// TIA Portal project "opc_pc-station" (V16)

(* hardware
DEVICE "S7-1200 station_1"  S7-1200 Station
   slot 0: "Rack_0"  S7-1200 Rack  Rack  V1.0
   slot 1: "1214dc"  CPU 1214C DC/DC/DC  6ES7 214-1AG40-0XB0  V4.4
DEVICE "PC station"  SIMATIC PC station
   slot 0: "PC station"  Rail  SIMATIC PC-Station  V1.0
      slot 125: "Stationmanager"  Station_Manager  V6.0.4
   slot 1: "IE general_1"  IE General  IE_CP  V8.2.0
   slot 2: "OPC Server_1"  OPC Server  OPC Server  V16.0.0
DEVICE "S7300/ET200M station_1"  S7-300 station
   slot 0: "Rail_0"  Rail  6ES7 390-1***0-0AA0
   slot 2: "314c"  CPU 314C-2 PN/DP  6ES7 314-6EH04-0AB0  V3.3
      slot 2: "PROFINET interface_1"  PN-IO
         slot 1: "Port_1"  Port
         slot 2: "Port_2"  Port
      slot 5: "DI 24/DO 16_1"  DI24/DO16
      slot 6: "AI 5/AO 2_1"  AI5/AO2
      slot 7: "Count_1"  Counter
      slot 8: "Positioning_1"  Positioning
DEVICE "S71500/ET200MP station_1"  S7-1500 station
   slot 0: "Rail_0"  Rack  6ES7 590-1***0-0AA0
   slot 1: "1511f"  CPU 1511F-1 PN  6ES7 511-1FK02-0AB0  V2.8
      slot 3: "CPU display_1"  6ES7591-1AA00-0AA0
      slot 32768: "1511f"  X1
         slot 32769: "Port_1"  X1 P1
         slot 32770: "Port_2"  X1 P2
      slot 34817: "Virtual CP interface port_1"  Virtual CP interface port  Virtual CP interface port
DEVICE "S7300/ET200M station_2"  S7-300 station
   slot 0: "Rail_0"  Rail  6ES7 390-1***0-0AA0
   slot 2: "314c_cp343"  CPU 314C-2 PN/DP  6ES7 314-6EH04-0AB0  V3.3
      slot 2: "PROFINET interface_1"  PN-IO
         slot 1: "Port_1"  Port
         slot 2: "Port_2"  Port
      slot 5: "DI 24/DO 16_1"  DI24/DO16
      slot 6: "AI 5/AO 2_1"  AI5/AO2
      slot 7: "Count_1"  Counter
      slot 8: "Positioning_1"  Positioning
   slot 4: "CP 343-1 Advanced-IT_1"  CP 343-1 ADVANCED-IT  6GK7 343-1GX31-0XE0  V3.0
DEVICE "S71500/ET200MP station_2"  S7-1500 station
   slot 0: "Rail_0"  Rack  6ES7 590-1***0-0AA0
   slot 1: "1511f_cp"  CPU 1511F-1 PN  6ES7 511-1FK02-0AB0  V2.8
      slot 3: "CPU display_1"  6ES7591-1AA00-0AA0
      slot 32768: "1511f"  X1
         slot 32769: "Port_1"  X1 P1
         slot 32770: "Port_2"  X1 P2
      slot 34817: "Virtual CP interface port_1"  Virtual CP interface port  Virtual CP interface port
   slot 2: "CP 1543-1_1"  CP 1543-1  6GK7 543-1AX00-0XE0  V2.2
DEVICE "S7-1200 station_2"  S7-1200 Station
   slot 0: "Rack_0"  S7-1200 Rack  Rack  V1.0
   slot 1: "1212fc_cp"  CPU 1212FC DC/DC/DC  6ES7 212-1AF40-0XB0  V4.4
   slot 101: "CP 1243-1"  CP 1243-1  6GK7 243-1BX30-0XE0  V3.2
      slot 0: "Telecontrol server"  Partner
      slot 0: "Inter-station communication"  Partner
*)

// ===== PLC "1214dc"  CPU 1214C DC/DC/DC =====

VAR_GLOBAL   // PLC tag table "Default tag table"
   "Tag_clock" AT %MW2 : Int;
   "Tag_Int" AT %MW4 : Int;
END_VAR

DATA_BLOCK "data_db"   // DB1
{ S7_Optimized_Access := 'TRUE' }
VERSION : 0.1
   VAR
      zm_array : Array[0..2] of Byte;
      zm_bool : Bool;
      zm_byte : Byte;
      zm_char : Char;
      zm_datetime_dtl : DTL;
      zm_dword : DWord;
      zm_int : Int;
      zm_real : Real;
      zm_string : String;
      zm_struct : Struct
         zm_struct_bool : Bool;
         zm_struct_byte : Byte;
      END_STRUCT;
   END_VAR
BEGIN
END_DATA_BLOCK

ORGANIZATION_BLOCK "Main"   // OB1, LAD, ProgramCycle
TITLE = "Main Program Sweep (Cycle)"
{ S7_Optimized_Access := 'TRUE' }
VERSION : 0.1
   VAR_INPUT
      Initial_Call : Bool;   // Initial call of this OB
      Remanence : Bool;   // =True, if remanent data are available
   END_VAR
BEGIN

REGION Network 1
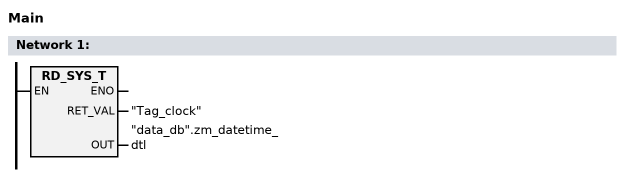
   "Tag_clock" := RD_SYS_T(OUT => "data_db".zm_datetime_dtl);
END_REGION
END_ORGANIZATION_BLOCK

// ===== PLC "314c"  CPU 314C-2 PN/DP =====

VAR_GLOBAL   // PLC tag table "Default tag table"
   "Tag_1" AT %MW0 : Int;
   "Tag_2" AT %M3.0 : Bool;
   "Tag_3" AT %MW4 : Word;
END_VAR

DATA_BLOCK "db_opc"   // DB1
{ S7_Optimized_Access := 'FALSE' }
VERSION : 0.1
   VAR
      zm_array : Array[0..2] of Byte;
      zm_bool : Bool;
      zm_byte : Byte;
      zm_char : Char;
      zm_datetime_rd_sys_t : Date_And_Time;
      zm_dword : DWord;
      zm_int : Int;
      zm_real : Real;
      zm_string : String;
      zm_struct : Struct
         zm_struct_bool : Bool;
         zm_struct_byte : Byte;
      END_STRUCT;
   END_VAR
BEGIN
END_DATA_BLOCK

ORGANIZATION_BLOCK "Main"   // OB1, LAD
TITLE = "Main Program Sweep (Cycle)"
{ S7_Optimized_Access := 'FALSE' }
VERSION : 0.1
   VAR_TEMP
      OB1_EV_CLASS : Byte;   // Bits 0-3 = 1 (Coming event), Bits 4-7 = 1 (Event class 1)
      OB1_SCAN_1 : Byte;   // 1 (Cold restart scan 1 of OB 1), 3 (Scan 2-n of OB 1)
      OB1_PRIORITY : Byte;   // Priority of OB Execution
      OB1_OB_NUMBR : Byte;   // 1 (Organization block 1, OB1)
      OB1_RESERVED_1 : Byte;   // Reserved for system
      OB1_RESERVED_2 : Byte;   // Reserved for system
      OB1_PREV_CYCLE : Int;   // Cycle time of previous OB1 scan (milliseconds)
      OB1_MIN_CYCLE : Int;   // Minimum cycle time of OB1 (milliseconds)
      OB1_MAX_CYCLE : Int;   // Maximum cycle time of OB1 (milliseconds)
      OB1_DATE_TIME : Date_And_Time;   // Date and time OB1 started
   END_VAR
BEGIN

REGION Network 1
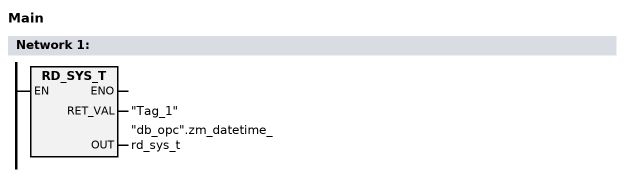
   "Tag_1" := RD_SYS_T(OUT => "db_opc".zm_datetime_rd_sys_t);
END_REGION
END_ORGANIZATION_BLOCK

// ===== PLC "1511f"  CPU 1511F-1 PN =====

VAR_GLOBAL   // PLC tag table "Default tag table"
   "Tag_1" AT %MW0 : Int;
END_VAR

DATA_BLOCK "data_db"   // DB1
{ S7_Optimized_Access := 'TRUE' }
VERSION : 0.1
   VAR
      zm_array : Array[0..2] of Byte;
      zm_bool : Bool;
      zm_byte : Byte;
      zm_char : Char;
      zm_datetime_dtl : DTL;
      zm_dword : DWord;
      zm_int : Int;
      zm_real : Real;
      zm_string : String;
      zm_struct : Struct
         zm_struct_bool : Bool;
         zm_struct_byte : Byte;
      END_STRUCT;
   END_VAR
BEGIN
END_DATA_BLOCK

ORGANIZATION_BLOCK "Main"   // OB1, LAD, ProgramCycle
TITLE = "Main Program Sweep (Cycle)"
{ S7_Optimized_Access := 'TRUE' }
VERSION : 0.1
   VAR_INPUT
      Initial_Call : Bool;   // Initial call of this OB
      Remanence : Bool;   // =True, if remanent data are available
   END_VAR
BEGIN

REGION Network 1
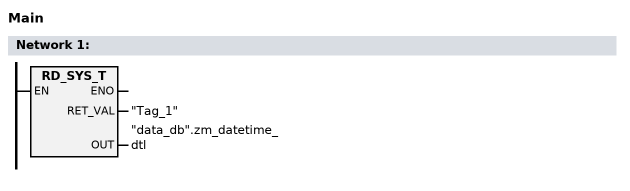
   "Tag_1" := RD_SYS_T(OUT => "data_db".zm_datetime_dtl);
END_REGION
END_ORGANIZATION_BLOCK

// ===== PLC "314c_cp343"  CPU 314C-2 PN/DP =====

VAR_GLOBAL   // PLC tag table "Default tag table"
   "Tag_1" AT %MW0 : Int;
   "Tag_2" AT %M3.0 : Bool;
   "Tag_3" AT %MW4 : Word;
END_VAR

DATA_BLOCK "db_opc"   // DB1
{ S7_Optimized_Access := 'FALSE' }
VERSION : 0.1
   VAR
      zm_array : Array[0..2] of Byte;
      zm_bool : Bool;
      zm_byte : Byte;
      zm_char : Char;
      zm_datetime_rd_sys_t : Date_And_Time;
      zm_dword : DWord;
      zm_int : Int;
      zm_real : Real;
      zm_string : String;
      zm_struct : Struct
         zm_struct_bool : Bool;
         zm_struct_byte : Byte;
      END_STRUCT;
   END_VAR
BEGIN
END_DATA_BLOCK

ORGANIZATION_BLOCK "Main"   // OB1, LAD
TITLE = "Main Program Sweep (Cycle)"
{ S7_Optimized_Access := 'FALSE' }
VERSION : 0.1
   VAR_TEMP
      OB1_EV_CLASS : Byte;   // Bits 0-3 = 1 (Coming event), Bits 4-7 = 1 (Event class 1)
      OB1_SCAN_1 : Byte;   // 1 (Cold restart scan 1 of OB 1), 3 (Scan 2-n of OB 1)
      OB1_PRIORITY : Byte;   // Priority of OB Execution
      OB1_OB_NUMBR : Byte;   // 1 (Organization block 1, OB1)
      OB1_RESERVED_1 : Byte;   // Reserved for system
      OB1_RESERVED_2 : Byte;   // Reserved for system
      OB1_PREV_CYCLE : Int;   // Cycle time of previous OB1 scan (milliseconds)
      OB1_MIN_CYCLE : Int;   // Minimum cycle time of OB1 (milliseconds)
      OB1_MAX_CYCLE : Int;   // Maximum cycle time of OB1 (milliseconds)
      OB1_DATE_TIME : Date_And_Time;   // Date and time OB1 started
   END_VAR
BEGIN

REGION Network 1
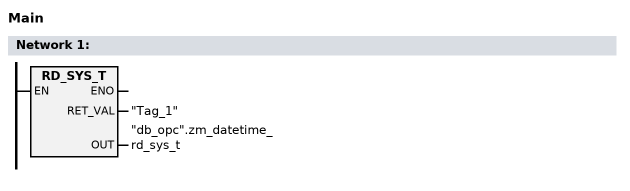
   "Tag_1" := RD_SYS_T(OUT => "db_opc".zm_datetime_rd_sys_t);
END_REGION
END_ORGANIZATION_BLOCK

// ===== PLC "1511f_cp"  CPU 1511F-1 PN =====

VAR_GLOBAL   // PLC tag table "Default tag table"
   "Tag_1" AT %MW0 : Int;
END_VAR

DATA_BLOCK "data_db"   // DB1
{ S7_Optimized_Access := 'TRUE' }
VERSION : 0.1
   VAR
      zm_array : Array[0..2] of Byte;
      zm_bool : Bool;
      zm_byte : Byte;
      zm_char : Char;
      zm_datetime_dtl : DTL;
      zm_dword : DWord;
      zm_int : Int;
      zm_real : Real;
      zm_string : String;
      zm_struct : Struct
         zm_struct_bool : Bool;
         zm_struct_byte : Byte;
      END_STRUCT;
   END_VAR
BEGIN
END_DATA_BLOCK

ORGANIZATION_BLOCK "Main"   // OB1, LAD, ProgramCycle
TITLE = "Main Program Sweep (Cycle)"
{ S7_Optimized_Access := 'TRUE' }
VERSION : 0.1
   VAR_INPUT
      Initial_Call : Bool;   // Initial call of this OB
      Remanence : Bool;   // =True, if remanent data are available
   END_VAR
BEGIN

REGION Network 1
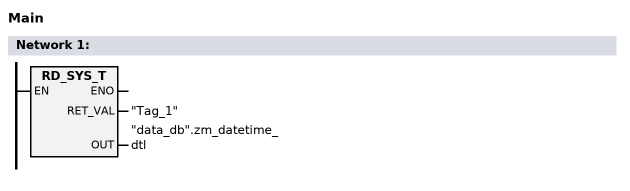
   "Tag_1" := RD_SYS_T(OUT => "data_db".zm_datetime_dtl);
END_REGION
END_ORGANIZATION_BLOCK

// ===== PLC "1212fc_cp"  CPU 1212FC DC/DC/DC =====

VAR_GLOBAL   // PLC tag table "Default tag table"
   "Tag_clock" AT %MW2 : Int;
   "Tag_Int" AT %MW4 : Int;
END_VAR

DATA_BLOCK "data_db"   // DB1
{ S7_Optimized_Access := 'TRUE' }
VERSION : 0.1
   VAR
      zm_array : Array[0..2] of Byte;
      zm_bool : Bool;
      zm_byte : Byte;
      zm_char : Char;
      zm_datetime_dtl : DTL;
      zm_dword : DWord;
      zm_int : Int;
      zm_real : Real;
      zm_string : String;
      zm_struct : Struct
         zm_struct_bool : Bool;
         zm_struct_byte : Byte;
      END_STRUCT;
   END_VAR
BEGIN
END_DATA_BLOCK

ORGANIZATION_BLOCK "Main"   // OB1, LAD, ProgramCycle
TITLE = "Main Program Sweep (Cycle)"
{ S7_Optimized_Access := 'TRUE' }
VERSION : 0.1
   VAR_INPUT
      Initial_Call : Bool;   // Initial call of this OB
      Remanence : Bool;   // =True, if remanent data are available
   END_VAR
BEGIN

REGION Network 1
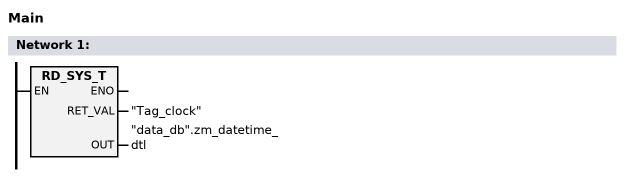
   "Tag_clock" := RD_SYS_T(OUT => "data_db".zm_datetime_dtl);
END_REGION
END_ORGANIZATION_BLOCK